(* Logix 5000 project; controller FV vendor 1 type 14 code 217 rev 31.11; software revision 31.00; part 22 of 63 *)
(* tags used below, declared in another part *)
   CheckTimeMask : INT;
   Delphi_Does_Eng_Func : BOOL;
   FR_FV29_AV04 : PlantItem;   // FV29_AV04
   FR_FV29_AV05 : PlantItem;   // FV29_AV05
   FR_FV29_AV06 : PlantItem;   // FV29_AV06
   FR_FV29_AV07 : PlantItem;   // FV29_AV07
   FR_N255 : INT[265];   // CHECKWORDS
   FR_VB2_AV01 : PlantItem;   // VB2_AV01
   FR_VB2_AV02 : PlantItem;   // VB2_AV02
   FR_VB2_AV03 : PlantItem;   // VB2_AV03
   FR_VB2_AV04 : PlantItem;   // VB2_AV04
   FR_VB2_AV05 : PlantItem;   // VB2_AV05
   FR_VB4_AV01 : PlantItem;   // VB4_AV01
   FR_VB4_AV02 : PlantItem;   // VB4_AV02
   FR_VB4_AV03 : PlantItem;   // VB4_AV03
   FR_VB4_AV04 : PlantItem;   // VB4_AV04
   TempChecktime : DINT;
(* FR_Common, continued *)

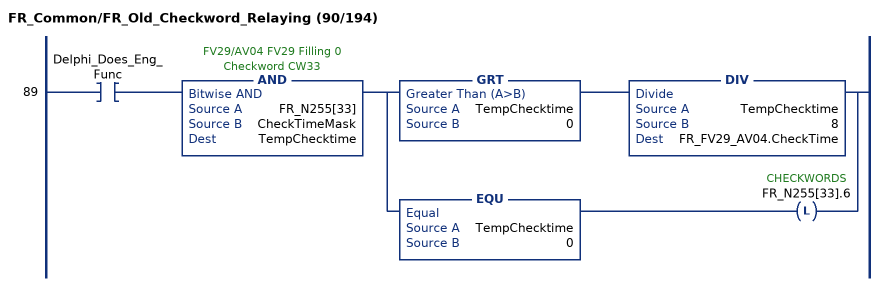
   [picture p394: FR_Common/FR_Old_Checkword_Relaying rungs 89-89]
   89: XIC(Delphi_Does_Eng_Func)AND(FR_N255[33],CheckTimeMask,TempChecktime)[GRT(TempChecktime,0) DIV(TempChecktime,8,FR_FV29_AV04.CheckTime) ,EQU(TempChecktime,0) OTL(FR_N255[33].6) ];
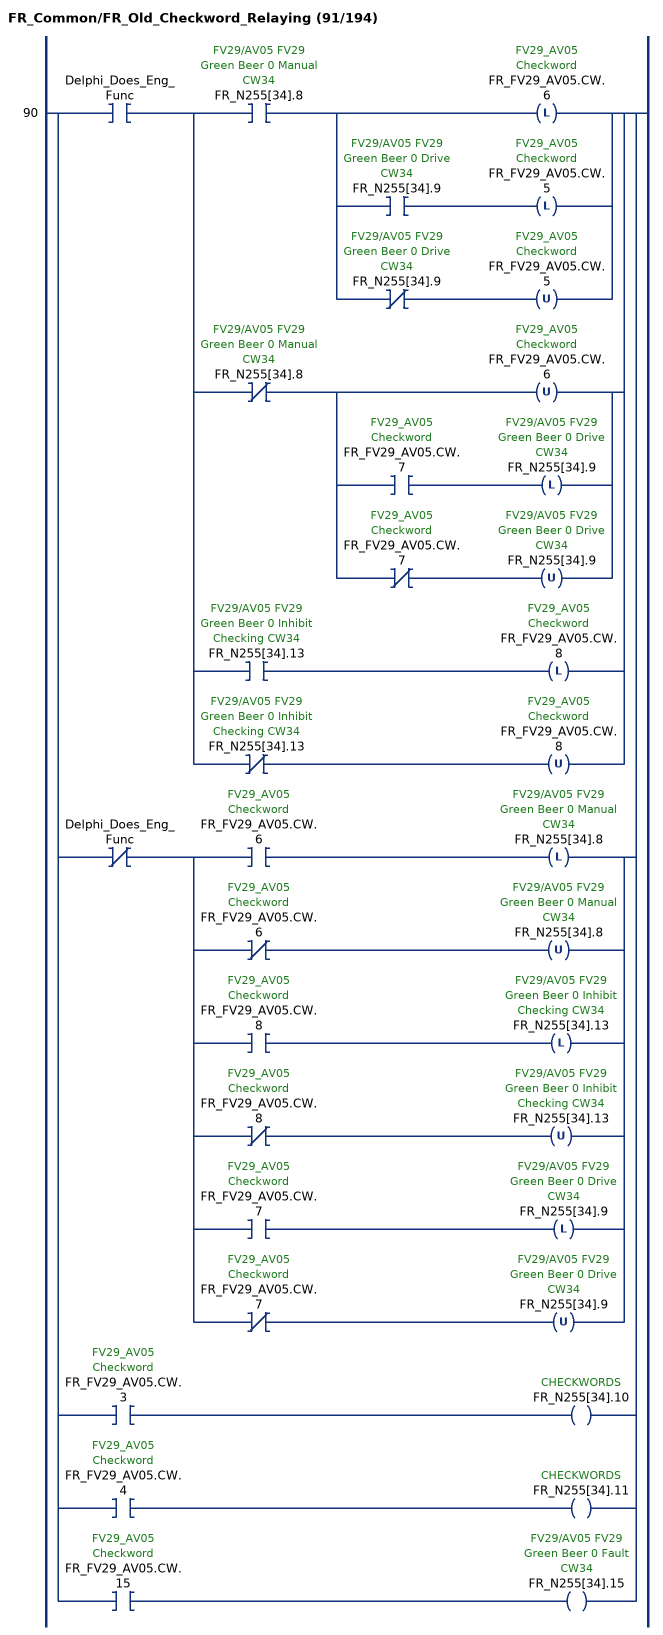
   90: [XIC(Delphi_Does_Eng_Func) [[XIC(FR_N255[34].8) [OTL(FR_FV29_AV05.CW.6) ,XIC(FR_N255[34].9) OTL(FR_FV29_AV05.CW.5) ,XIO(FR_N255[34].9) OTU(FR_FV29_AV05.CW.5) ] ,XIO(FR_N255[34].8) [OTU(FR_FV29_AV05.CW.6) ,[XIC(FR_FV29_AV05.CW.7) OTL(FR_N255[34].9) ,XIO(FR_FV29_AV05.CW.7) OTU(FR_N255[34].9) ] ] ] ,[XIC(FR_N255[34].13) OTL(FR_FV29_AV05.CW.8) ,XIO(FR_N255[34].13) OTU(FR_FV29_AV05.CW.8) ] ] ,XIO(Delphi_Does_Eng_Func) [[XIC(FR_FV29_AV05.CW.6) OTL(FR_N255[34].8) ,XIO(FR_FV29_AV05.CW.6) OTU(FR_N255[34].8) ] ,[XIC(FR_FV29_AV05.CW.8) OTL(FR_N255[34].13) ,XIO(FR_FV29_AV05.CW.8) OTU(FR_N255[34].13) ] ,[XIC(FR_FV29_AV05.CW.7) OTL(FR_N255[34].9) ,XIO(FR_FV29_AV05.CW.7) OTU(FR_N255[34].9) ] ] ,XIC(FR_FV29_AV05.CW.3) OTE(FR_N255[34].10) ,XIC(FR_FV29_AV05.CW.4) OTE(FR_N255[34].11) ,XIC(FR_FV29_AV05.CW.15) OTE(FR_N255[34].15) ];
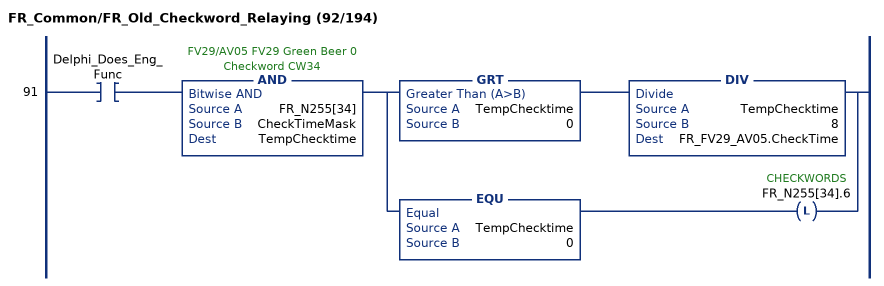
   91: XIC(Delphi_Does_Eng_Func)AND(FR_N255[34],CheckTimeMask,TempChecktime)[GRT(TempChecktime,0) DIV(TempChecktime,8,FR_FV29_AV05.CheckTime) ,EQU(TempChecktime,0) OTL(FR_N255[34].6) ];
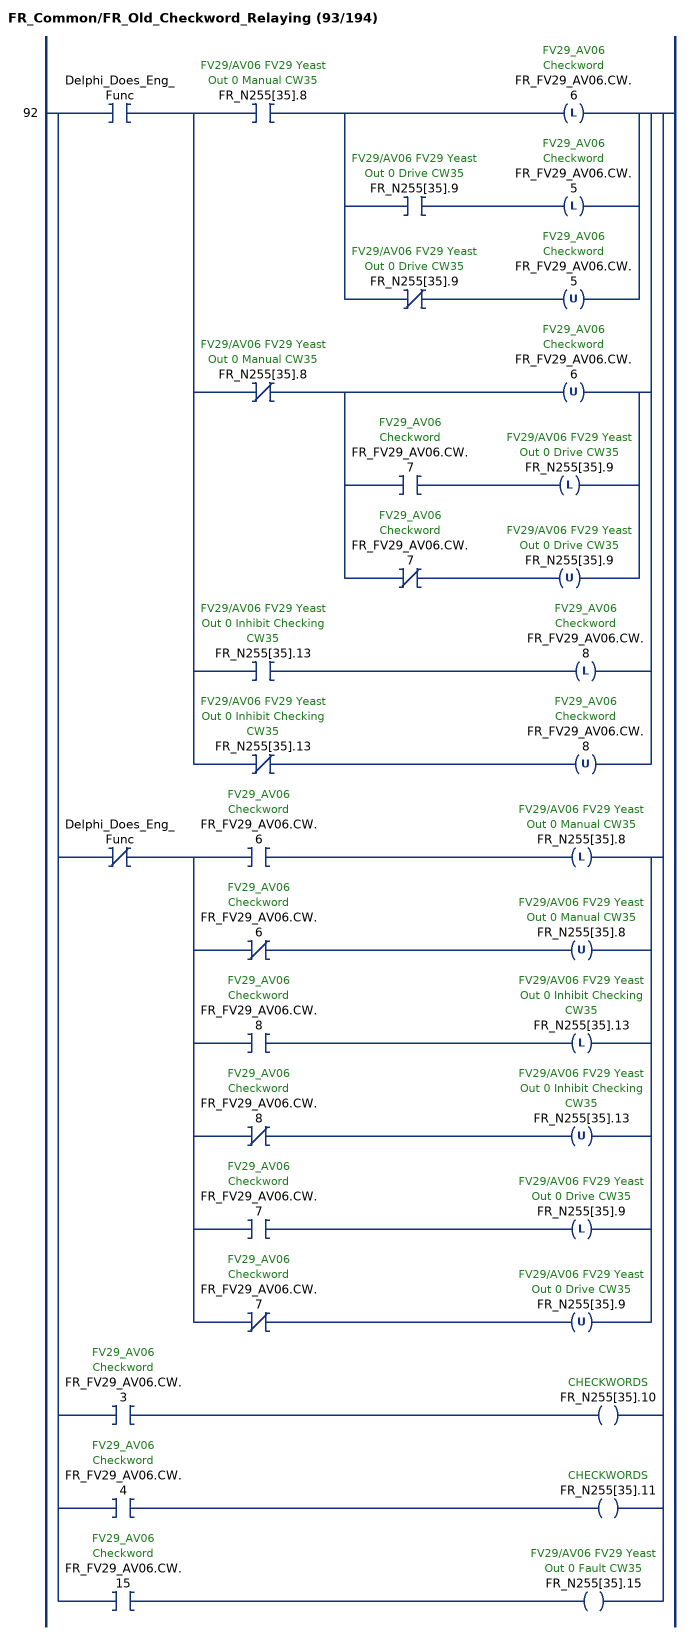
   92: [XIC(Delphi_Does_Eng_Func) [[XIC(FR_N255[35].8) [OTL(FR_FV29_AV06.CW.6) ,XIC(FR_N255[35].9) OTL(FR_FV29_AV06.CW.5) ,XIO(FR_N255[35].9) OTU(FR_FV29_AV06.CW.5) ] ,XIO(FR_N255[35].8) [OTU(FR_FV29_AV06.CW.6) ,[XIC(FR_FV29_AV06.CW.7) OTL(FR_N255[35].9) ,XIO(FR_FV29_AV06.CW.7) OTU(FR_N255[35].9) ] ] ] ,[XIC(FR_N255[35].13) OTL(FR_FV29_AV06.CW.8) ,XIO(FR_N255[35].13) OTU(FR_FV29_AV06.CW.8) ] ] ,XIO(Delphi_Does_Eng_Func) [[XIC(FR_FV29_AV06.CW.6) OTL(FR_N255[35].8) ,XIO(FR_FV29_AV06.CW.6) OTU(FR_N255[35].8) ] ,[XIC(FR_FV29_AV06.CW.8) OTL(FR_N255[35].13) ,XIO(FR_FV29_AV06.CW.8) OTU(FR_N255[35].13) ] ,[XIC(FR_FV29_AV06.CW.7) OTL(FR_N255[35].9) ,XIO(FR_FV29_AV06.CW.7) OTU(FR_N255[35].9) ] ] ,XIC(FR_FV29_AV06.CW.3) OTE(FR_N255[35].10) ,XIC(FR_FV29_AV06.CW.4) OTE(FR_N255[35].11) ,XIC(FR_FV29_AV06.CW.15) OTE(FR_N255[35].15) ];
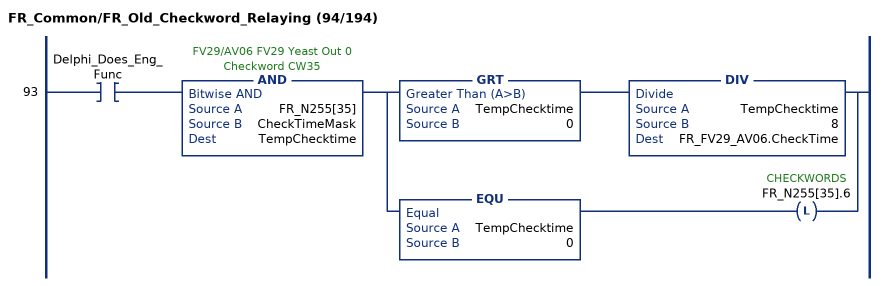
   93: XIC(Delphi_Does_Eng_Func)AND(FR_N255[35],CheckTimeMask,TempChecktime)[GRT(TempChecktime,0) DIV(TempChecktime,8,FR_FV29_AV06.CheckTime) ,EQU(TempChecktime,0) OTL(FR_N255[35].6) ];
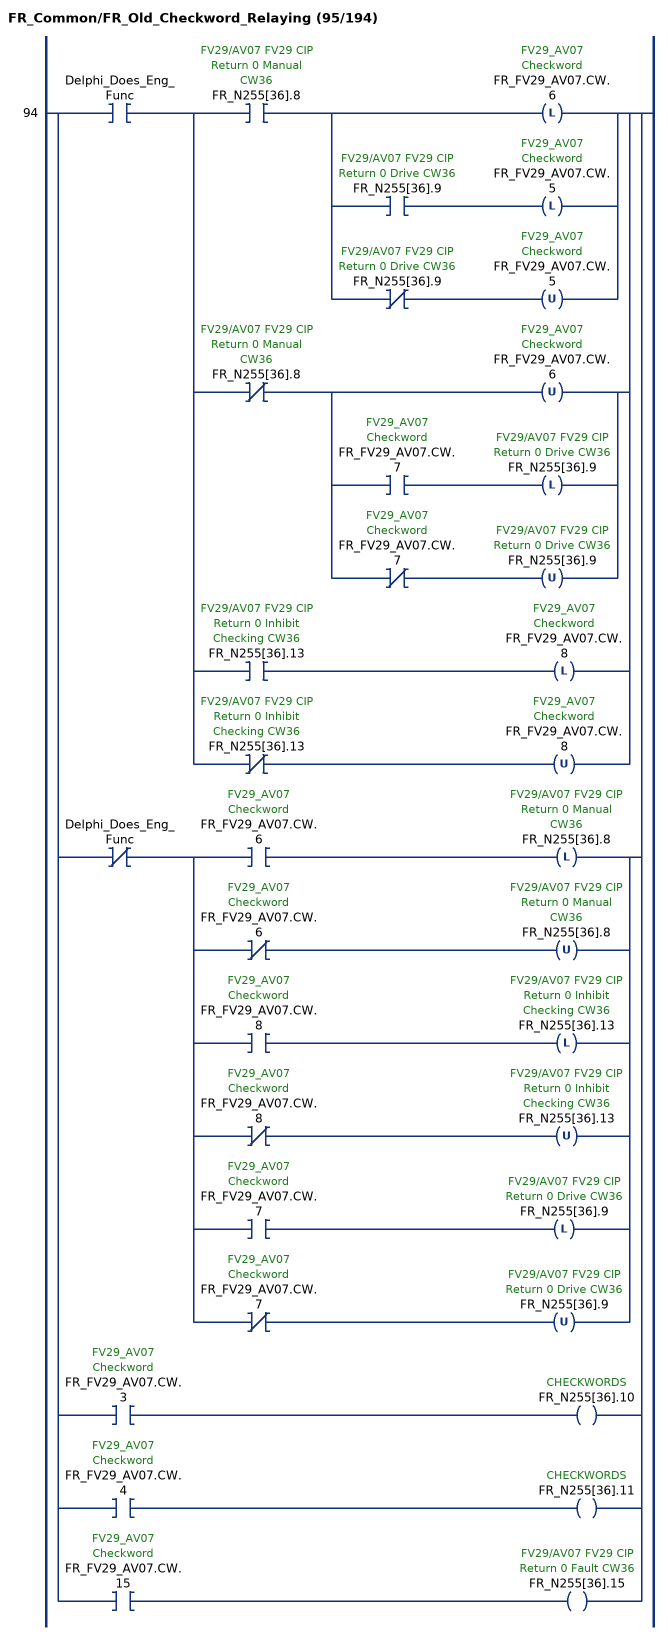
   94: [XIC(Delphi_Does_Eng_Func) [[XIC(FR_N255[36].8) [OTL(FR_FV29_AV07.CW.6) ,XIC(FR_N255[36].9) OTL(FR_FV29_AV07.CW.5) ,XIO(FR_N255[36].9) OTU(FR_FV29_AV07.CW.5) ] ,XIO(FR_N255[36].8) [OTU(FR_FV29_AV07.CW.6) ,[XIC(FR_FV29_AV07.CW.7) OTL(FR_N255[36].9) ,XIO(FR_FV29_AV07.CW.7) OTU(FR_N255[36].9) ] ] ] ,[XIC(FR_N255[36].13) OTL(FR_FV29_AV07.CW.8) ,XIO(FR_N255[36].13) OTU(FR_FV29_AV07.CW.8) ] ] ,XIO(Delphi_Does_Eng_Func) [[XIC(FR_FV29_AV07.CW.6) OTL(FR_N255[36].8) ,XIO(FR_FV29_AV07.CW.6) OTU(FR_N255[36].8) ] ,[XIC(FR_FV29_AV07.CW.8) OTL(FR_N255[36].13) ,XIO(FR_FV29_AV07.CW.8) OTU(FR_N255[36].13) ] ,[XIC(FR_FV29_AV07.CW.7) OTL(FR_N255[36].9) ,XIO(FR_FV29_AV07.CW.7) OTU(FR_N255[36].9) ] ] ,XIC(FR_FV29_AV07.CW.3) OTE(FR_N255[36].10) ,XIC(FR_FV29_AV07.CW.4) OTE(FR_N255[36].11) ,XIC(FR_FV29_AV07.CW.15) OTE(FR_N255[36].15) ];
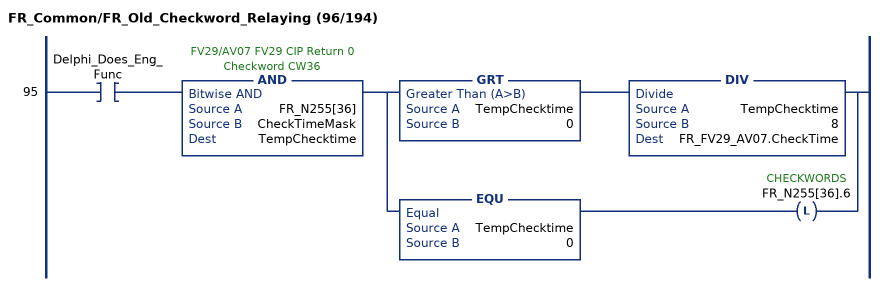
   95: XIC(Delphi_Does_Eng_Func)AND(FR_N255[36],CheckTimeMask,TempChecktime)[GRT(TempChecktime,0) DIV(TempChecktime,8,FR_FV29_AV07.CheckTime) ,EQU(TempChecktime,0) OTL(FR_N255[36].6) ];
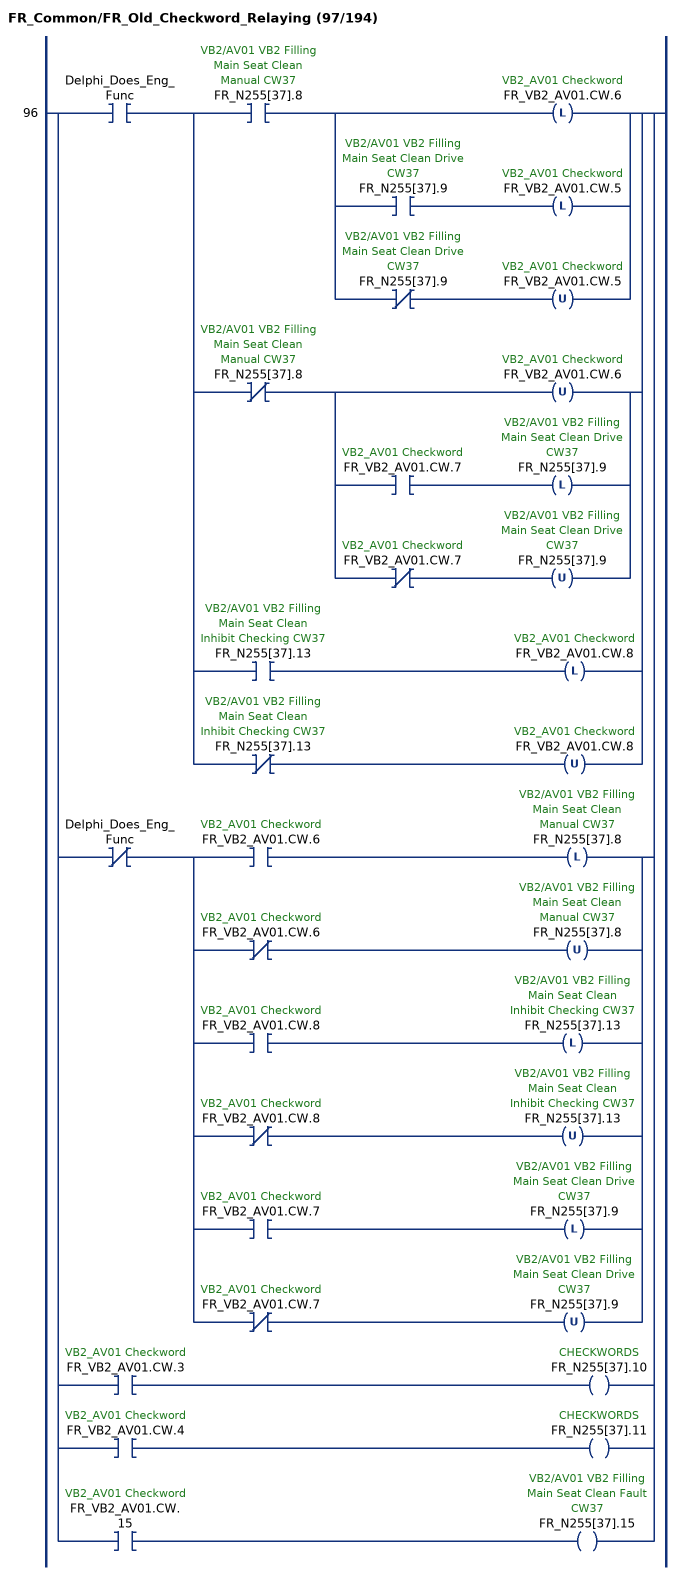
   96: [XIC(Delphi_Does_Eng_Func) [[XIC(FR_N255[37].8) [OTL(FR_VB2_AV01.CW.6) ,XIC(FR_N255[37].9) OTL(FR_VB2_AV01.CW.5) ,XIO(FR_N255[37].9) OTU(FR_VB2_AV01.CW.5) ] ,XIO(FR_N255[37].8) [OTU(FR_VB2_AV01.CW.6) ,[XIC(FR_VB2_AV01.CW.7) OTL(FR_N255[37].9) ,XIO(FR_VB2_AV01.CW.7) OTU(FR_N255[37].9) ] ] ] ,[XIC(FR_N255[37].13) OTL(FR_VB2_AV01.CW.8) ,XIO(FR_N255[37].13) OTU(FR_VB2_AV01.CW.8) ] ] ,XIO(Delphi_Does_Eng_Func) [[XIC(FR_VB2_AV01.CW.6) OTL(FR_N255[37].8) ,XIO(FR_VB2_AV01.CW.6) OTU(FR_N255[37].8) ] ,[XIC(FR_VB2_AV01.CW.8) OTL(FR_N255[37].13) ,XIO(FR_VB2_AV01.CW.8) OTU(FR_N255[37].13) ] ,[XIC(FR_VB2_AV01.CW.7) OTL(FR_N255[37].9) ,XIO(FR_VB2_AV01.CW.7) OTU(FR_N255[37].9) ] ] ,XIC(FR_VB2_AV01.CW.3) OTE(FR_N255[37].10) ,XIC(FR_VB2_AV01.CW.4) OTE(FR_N255[37].11) ,XIC(FR_VB2_AV01.CW.15) OTE(FR_N255[37].15) ];
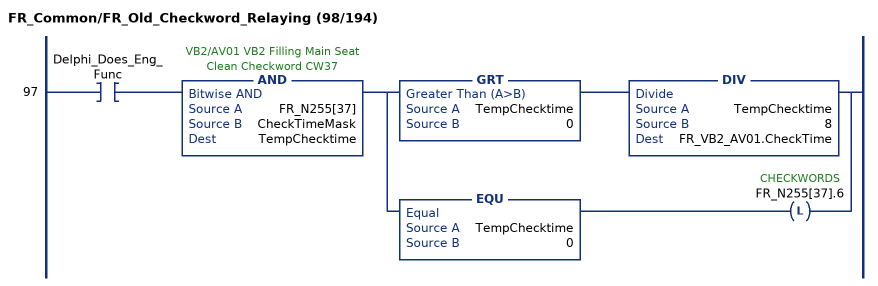
   97: XIC(Delphi_Does_Eng_Func)AND(FR_N255[37],CheckTimeMask,TempChecktime)[GRT(TempChecktime,0) DIV(TempChecktime,8,FR_VB2_AV01.CheckTime) ,EQU(TempChecktime,0) OTL(FR_N255[37].6) ];
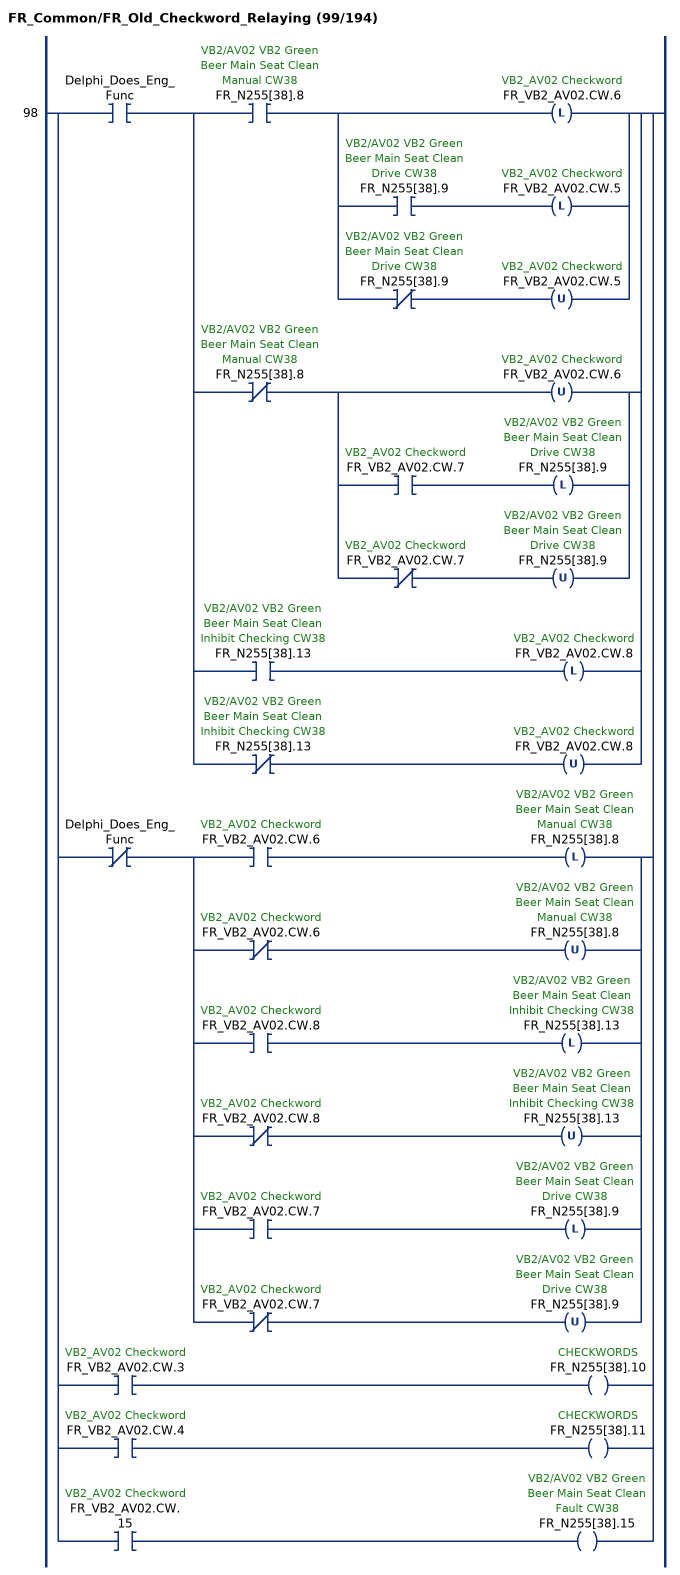
   98: [XIC(Delphi_Does_Eng_Func) [[XIC(FR_N255[38].8) [OTL(FR_VB2_AV02.CW.6) ,XIC(FR_N255[38].9) OTL(FR_VB2_AV02.CW.5) ,XIO(FR_N255[38].9) OTU(FR_VB2_AV02.CW.5) ] ,XIO(FR_N255[38].8) [OTU(FR_VB2_AV02.CW.6) ,[XIC(FR_VB2_AV02.CW.7) OTL(FR_N255[38].9) ,XIO(FR_VB2_AV02.CW.7) OTU(FR_N255[38].9) ] ] ] ,[XIC(FR_N255[38].13) OTL(FR_VB2_AV02.CW.8) ,XIO(FR_N255[38].13) OTU(FR_VB2_AV02.CW.8) ] ] ,XIO(Delphi_Does_Eng_Func) [[XIC(FR_VB2_AV02.CW.6) OTL(FR_N255[38].8) ,XIO(FR_VB2_AV02.CW.6) OTU(FR_N255[38].8) ] ,[XIC(FR_VB2_AV02.CW.8) OTL(FR_N255[38].13) ,XIO(FR_VB2_AV02.CW.8) OTU(FR_N255[38].13) ] ,[XIC(FR_VB2_AV02.CW.7) OTL(FR_N255[38].9) ,XIO(FR_VB2_AV02.CW.7) OTU(FR_N255[38].9) ] ] ,XIC(FR_VB2_AV02.CW.3) OTE(FR_N255[38].10) ,XIC(FR_VB2_AV02.CW.4) OTE(FR_N255[38].11) ,XIC(FR_VB2_AV02.CW.15) OTE(FR_N255[38].15) ];
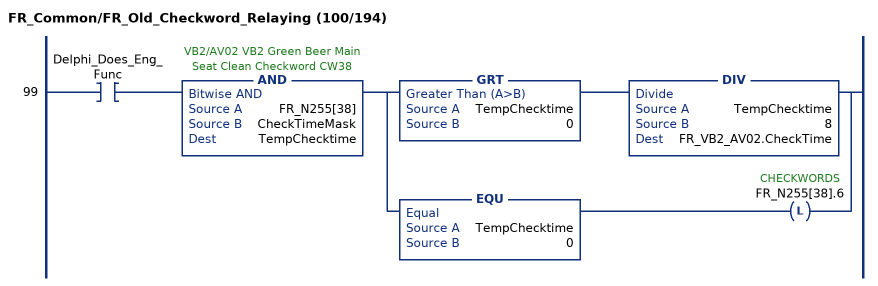
   99: XIC(Delphi_Does_Eng_Func)AND(FR_N255[38],CheckTimeMask,TempChecktime)[GRT(TempChecktime,0) DIV(TempChecktime,8,FR_VB2_AV02.CheckTime) ,EQU(TempChecktime,0) OTL(FR_N255[38].6) ];
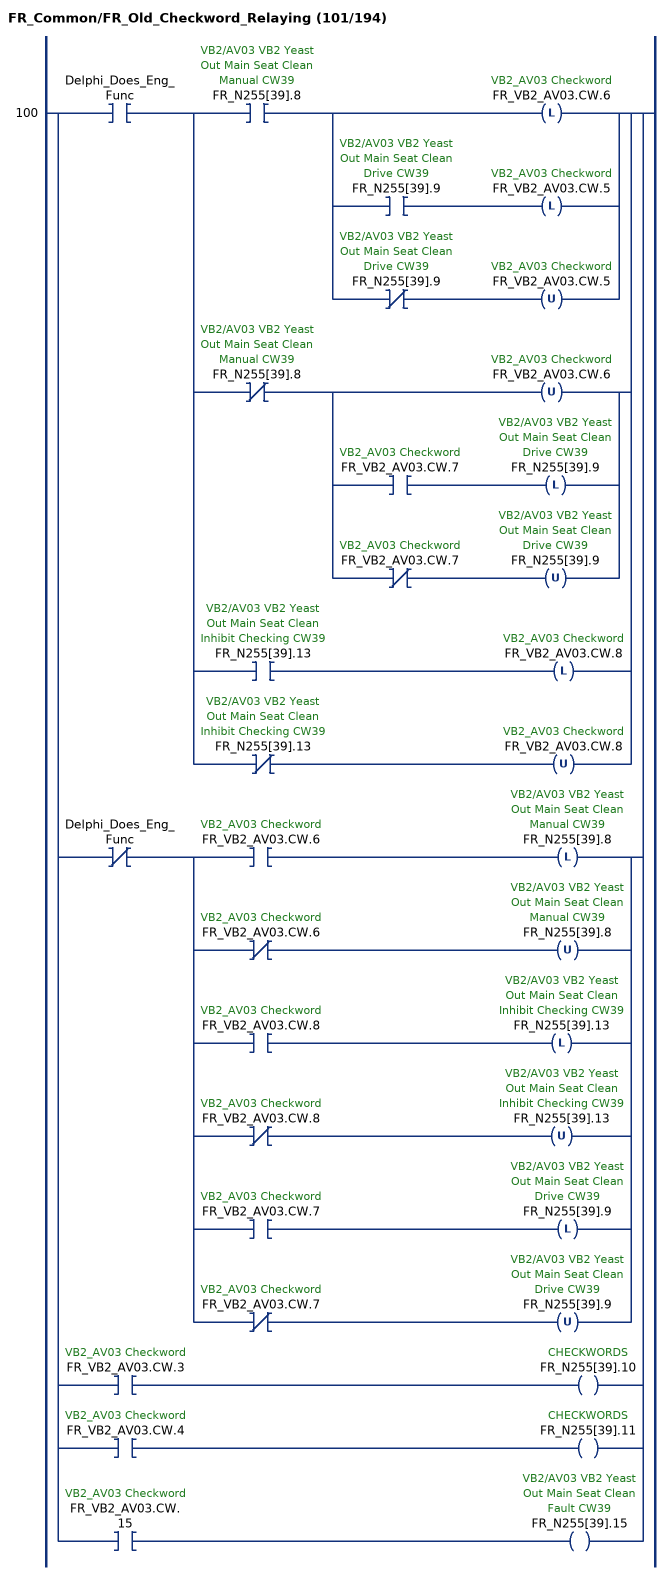
   100: [XIC(Delphi_Does_Eng_Func) [[XIC(FR_N255[39].8) [OTL(FR_VB2_AV03.CW.6) ,XIC(FR_N255[39].9) OTL(FR_VB2_AV03.CW.5) ,XIO(FR_N255[39].9) OTU(FR_VB2_AV03.CW.5) ] ,XIO(FR_N255[39].8) [OTU(FR_VB2_AV03.CW.6) ,[XIC(FR_VB2_AV03.CW.7) OTL(FR_N255[39].9) ,XIO(FR_VB2_AV03.CW.7) OTU(FR_N255[39].9) ] ] ] ,[XIC(FR_N255[39].13) OTL(FR_VB2_AV03.CW.8) ,XIO(FR_N255[39].13) OTU(FR_VB2_AV03.CW.8) ] ] ,XIO(Delphi_Does_Eng_Func) [[XIC(FR_VB2_AV03.CW.6) OTL(FR_N255[39].8) ,XIO(FR_VB2_AV03.CW.6) OTU(FR_N255[39].8) ] ,[XIC(FR_VB2_AV03.CW.8) OTL(FR_N255[39].13) ,XIO(FR_VB2_AV03.CW.8) OTU(FR_N255[39].13) ] ,[XIC(FR_VB2_AV03.CW.7) OTL(FR_N255[39].9) ,XIO(FR_VB2_AV03.CW.7) OTU(FR_N255[39].9) ] ] ,XIC(FR_VB2_AV03.CW.3) OTE(FR_N255[39].10) ,XIC(FR_VB2_AV03.CW.4) OTE(FR_N255[39].11) ,XIC(FR_VB2_AV03.CW.15) OTE(FR_N255[39].15) ];
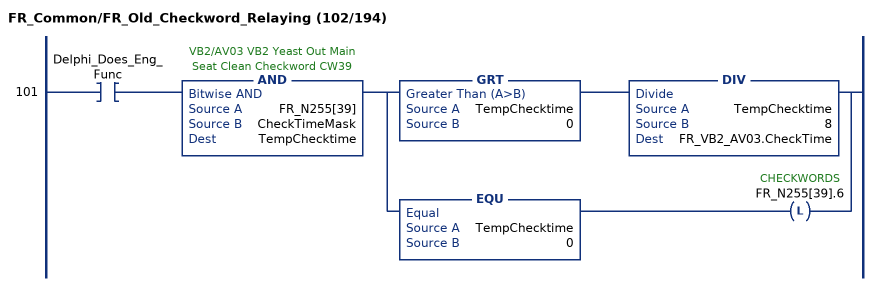
   101: XIC(Delphi_Does_Eng_Func)AND(FR_N255[39],CheckTimeMask,TempChecktime)[GRT(TempChecktime,0) DIV(TempChecktime,8,FR_VB2_AV03.CheckTime) ,EQU(TempChecktime,0) OTL(FR_N255[39].6) ];
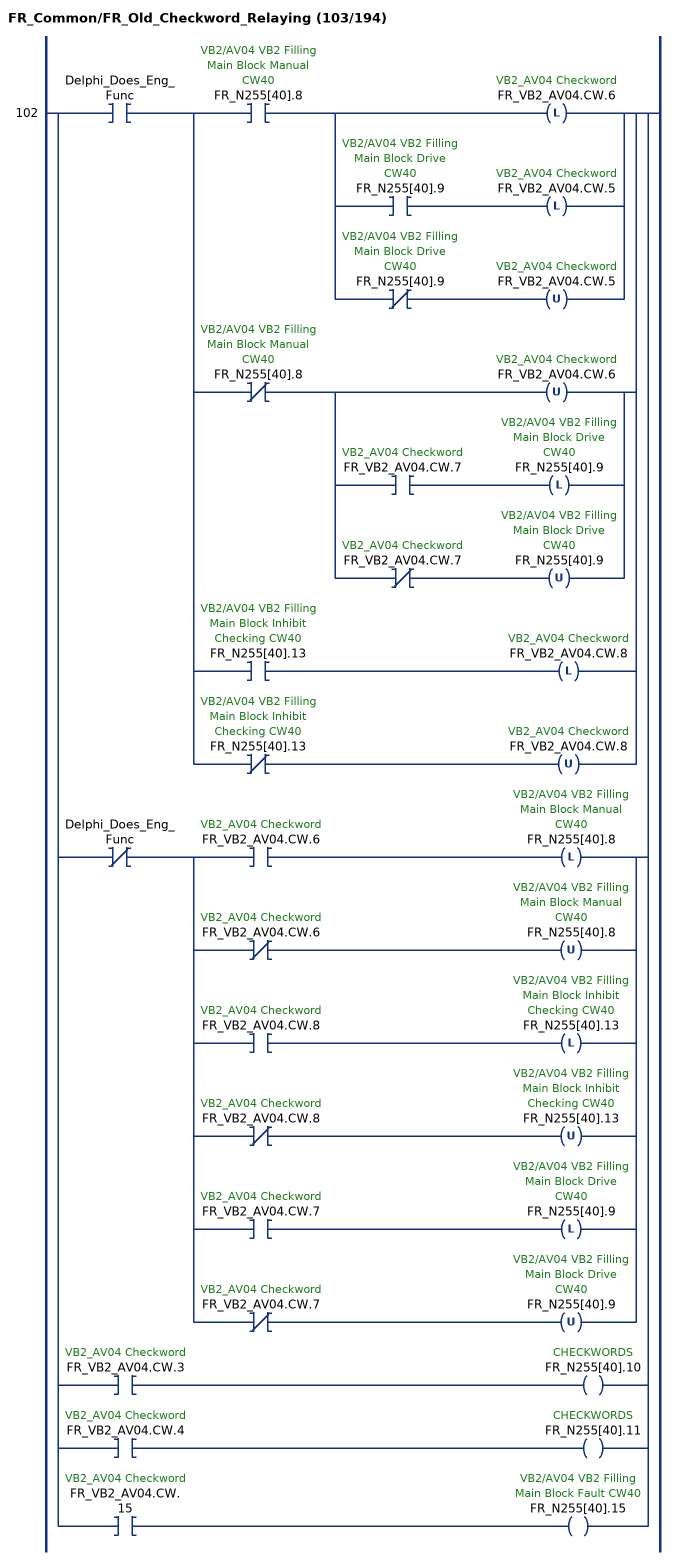
   102: [XIC(Delphi_Does_Eng_Func) [[XIC(FR_N255[40].8) [OTL(FR_VB2_AV04.CW.6) ,XIC(FR_N255[40].9) OTL(FR_VB2_AV04.CW.5) ,XIO(FR_N255[40].9) OTU(FR_VB2_AV04.CW.5) ] ,XIO(FR_N255[40].8) [OTU(FR_VB2_AV04.CW.6) ,[XIC(FR_VB2_AV04.CW.7) OTL(FR_N255[40].9) ,XIO(FR_VB2_AV04.CW.7) OTU(FR_N255[40].9) ] ] ] ,[XIC(FR_N255[40].13) OTL(FR_VB2_AV04.CW.8) ,XIO(FR_N255[40].13) OTU(FR_VB2_AV04.CW.8) ] ] ,XIO(Delphi_Does_Eng_Func) [[XIC(FR_VB2_AV04.CW.6) OTL(FR_N255[40].8) ,XIO(FR_VB2_AV04.CW.6) OTU(FR_N255[40].8) ] ,[XIC(FR_VB2_AV04.CW.8) OTL(FR_N255[40].13) ,XIO(FR_VB2_AV04.CW.8) OTU(FR_N255[40].13) ] ,[XIC(FR_VB2_AV04.CW.7) OTL(FR_N255[40].9) ,XIO(FR_VB2_AV04.CW.7) OTU(FR_N255[40].9) ] ] ,XIC(FR_VB2_AV04.CW.3) OTE(FR_N255[40].10) ,XIC(FR_VB2_AV04.CW.4) OTE(FR_N255[40].11) ,XIC(FR_VB2_AV04.CW.15) OTE(FR_N255[40].15) ];
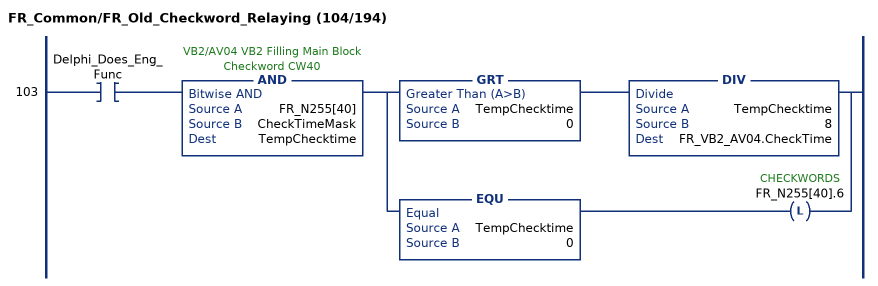
   103: XIC(Delphi_Does_Eng_Func)AND(FR_N255[40],CheckTimeMask,TempChecktime)[GRT(TempChecktime,0) DIV(TempChecktime,8,FR_VB2_AV04.CheckTime) ,EQU(TempChecktime,0) OTL(FR_N255[40].6) ];
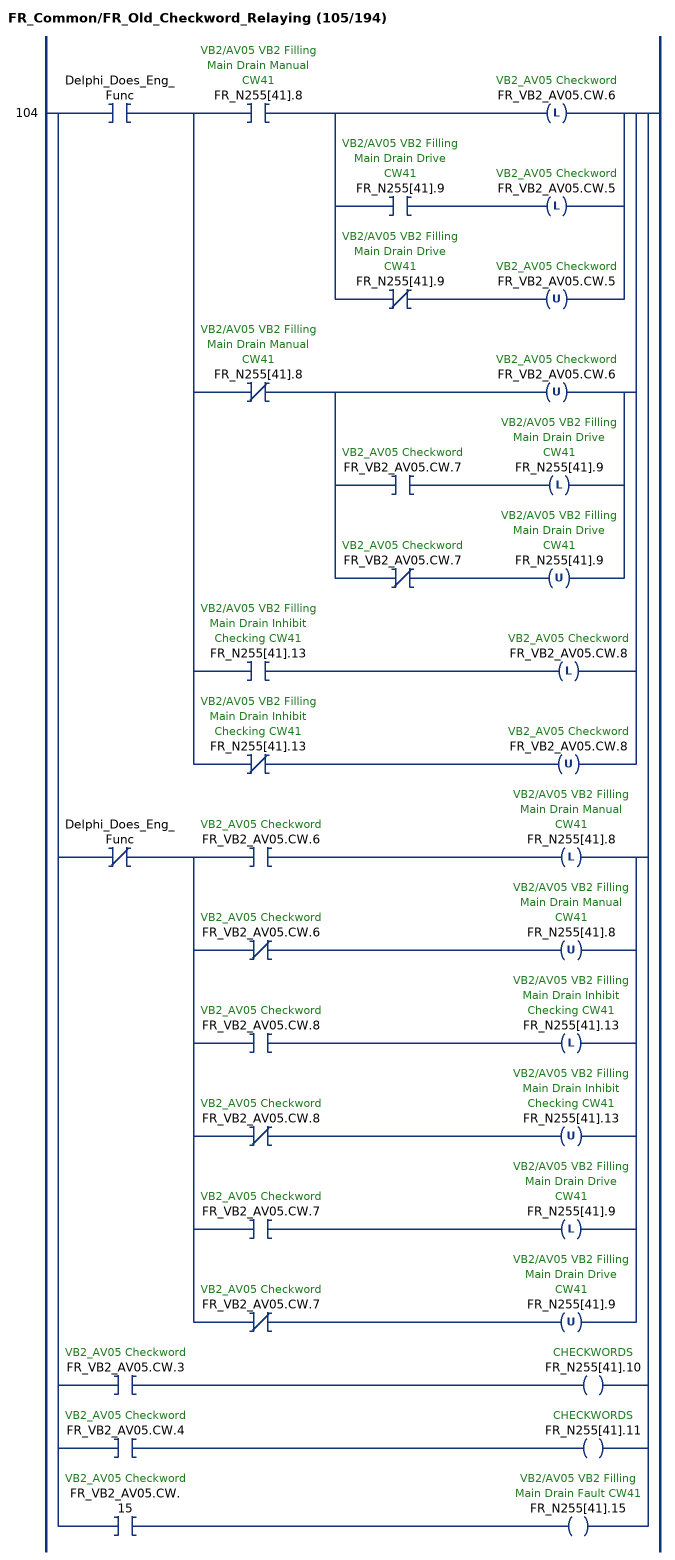
   104: [XIC(Delphi_Does_Eng_Func) [[XIC(FR_N255[41].8) [OTL(FR_VB2_AV05.CW.6) ,XIC(FR_N255[41].9) OTL(FR_VB2_AV05.CW.5) ,XIO(FR_N255[41].9) OTU(FR_VB2_AV05.CW.5) ] ,XIO(FR_N255[41].8) [OTU(FR_VB2_AV05.CW.6) ,[XIC(FR_VB2_AV05.CW.7) OTL(FR_N255[41].9) ,XIO(FR_VB2_AV05.CW.7) OTU(FR_N255[41].9) ] ] ] ,[XIC(FR_N255[41].13) OTL(FR_VB2_AV05.CW.8) ,XIO(FR_N255[41].13) OTU(FR_VB2_AV05.CW.8) ] ] ,XIO(Delphi_Does_Eng_Func) [[XIC(FR_VB2_AV05.CW.6) OTL(FR_N255[41].8) ,XIO(FR_VB2_AV05.CW.6) OTU(FR_N255[41].8) ] ,[XIC(FR_VB2_AV05.CW.8) OTL(FR_N255[41].13) ,XIO(FR_VB2_AV05.CW.8) OTU(FR_N255[41].13) ] ,[XIC(FR_VB2_AV05.CW.7) OTL(FR_N255[41].9) ,XIO(FR_VB2_AV05.CW.7) OTU(FR_N255[41].9) ] ] ,XIC(FR_VB2_AV05.CW.3) OTE(FR_N255[41].10) ,XIC(FR_VB2_AV05.CW.4) OTE(FR_N255[41].11) ,XIC(FR_VB2_AV05.CW.15) OTE(FR_N255[41].15) ];
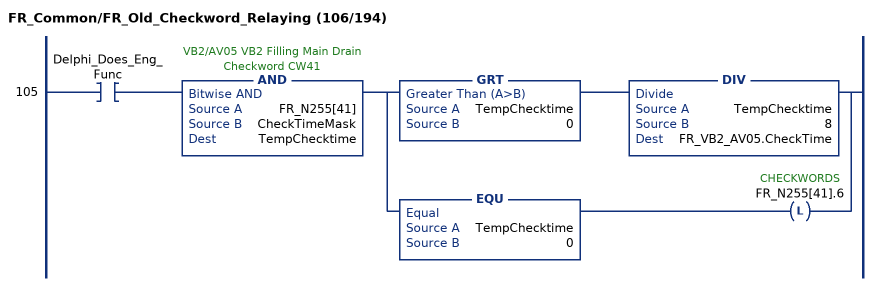
   105: XIC(Delphi_Does_Eng_Func)AND(FR_N255[41],CheckTimeMask,TempChecktime)[GRT(TempChecktime,0) DIV(TempChecktime,8,FR_VB2_AV05.CheckTime) ,EQU(TempChecktime,0) OTL(FR_N255[41].6) ];
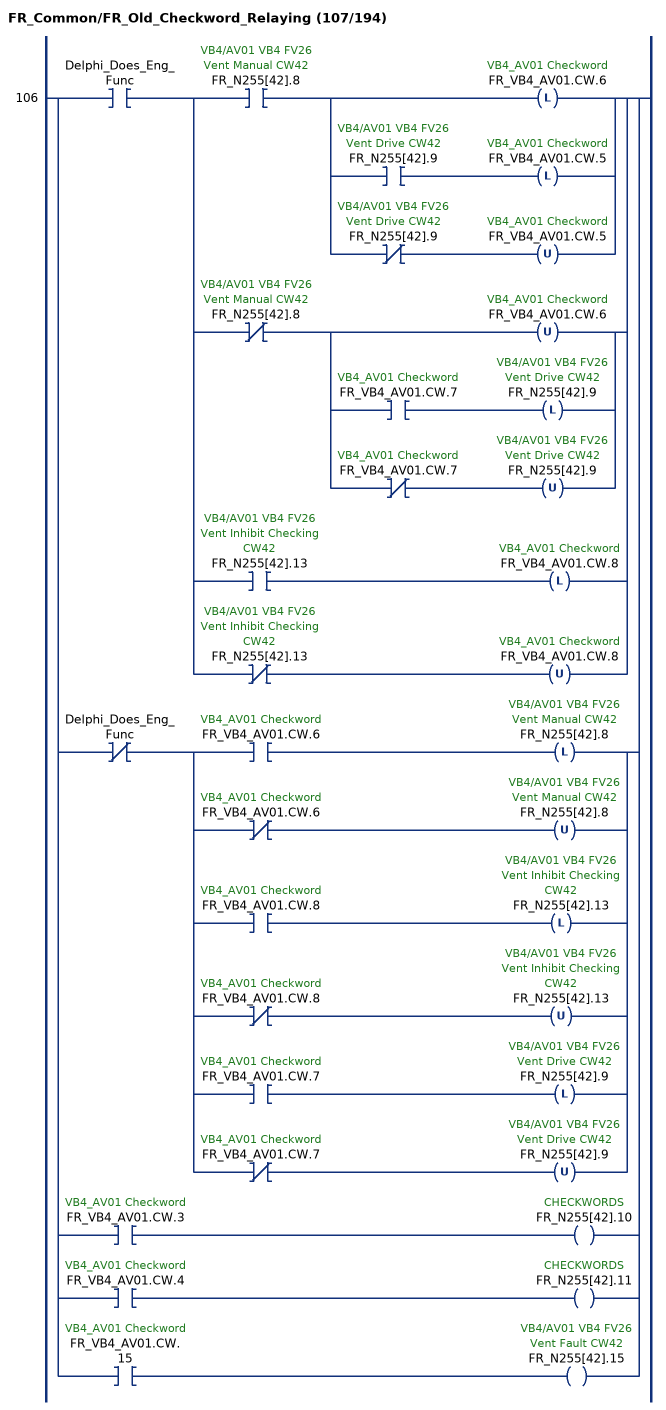
   106: [XIC(Delphi_Does_Eng_Func) [[XIC(FR_N255[42].8) [OTL(FR_VB4_AV01.CW.6) ,XIC(FR_N255[42].9) OTL(FR_VB4_AV01.CW.5) ,XIO(FR_N255[42].9) OTU(FR_VB4_AV01.CW.5) ] ,XIO(FR_N255[42].8) [OTU(FR_VB4_AV01.CW.6) ,[XIC(FR_VB4_AV01.CW.7) OTL(FR_N255[42].9) ,XIO(FR_VB4_AV01.CW.7) OTU(FR_N255[42].9) ] ] ] ,[XIC(FR_N255[42].13) OTL(FR_VB4_AV01.CW.8) ,XIO(FR_N255[42].13) OTU(FR_VB4_AV01.CW.8) ] ] ,XIO(Delphi_Does_Eng_Func) [[XIC(FR_VB4_AV01.CW.6) OTL(FR_N255[42].8) ,XIO(FR_VB4_AV01.CW.6) OTU(FR_N255[42].8) ] ,[XIC(FR_VB4_AV01.CW.8) OTL(FR_N255[42].13) ,XIO(FR_VB4_AV01.CW.8) OTU(FR_N255[42].13) ] ,[XIC(FR_VB4_AV01.CW.7) OTL(FR_N255[42].9) ,XIO(FR_VB4_AV01.CW.7) OTU(FR_N255[42].9) ] ] ,XIC(FR_VB4_AV01.CW.3) OTE(FR_N255[42].10) ,XIC(FR_VB4_AV01.CW.4) OTE(FR_N255[42].11) ,XIC(FR_VB4_AV01.CW.15) OTE(FR_N255[42].15) ];
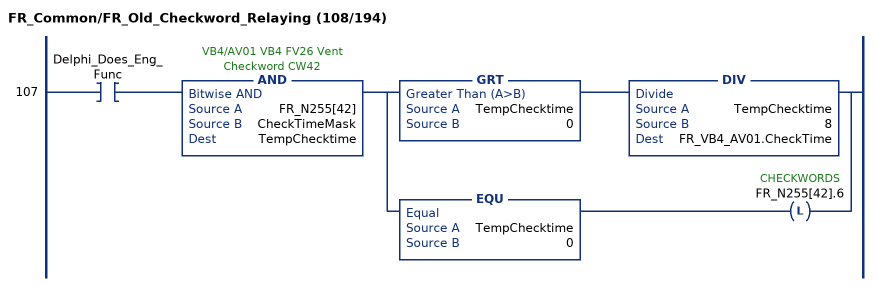
   107: XIC(Delphi_Does_Eng_Func)AND(FR_N255[42],CheckTimeMask,TempChecktime)[GRT(TempChecktime,0) DIV(TempChecktime,8,FR_VB4_AV01.CheckTime) ,EQU(TempChecktime,0) OTL(FR_N255[42].6) ];
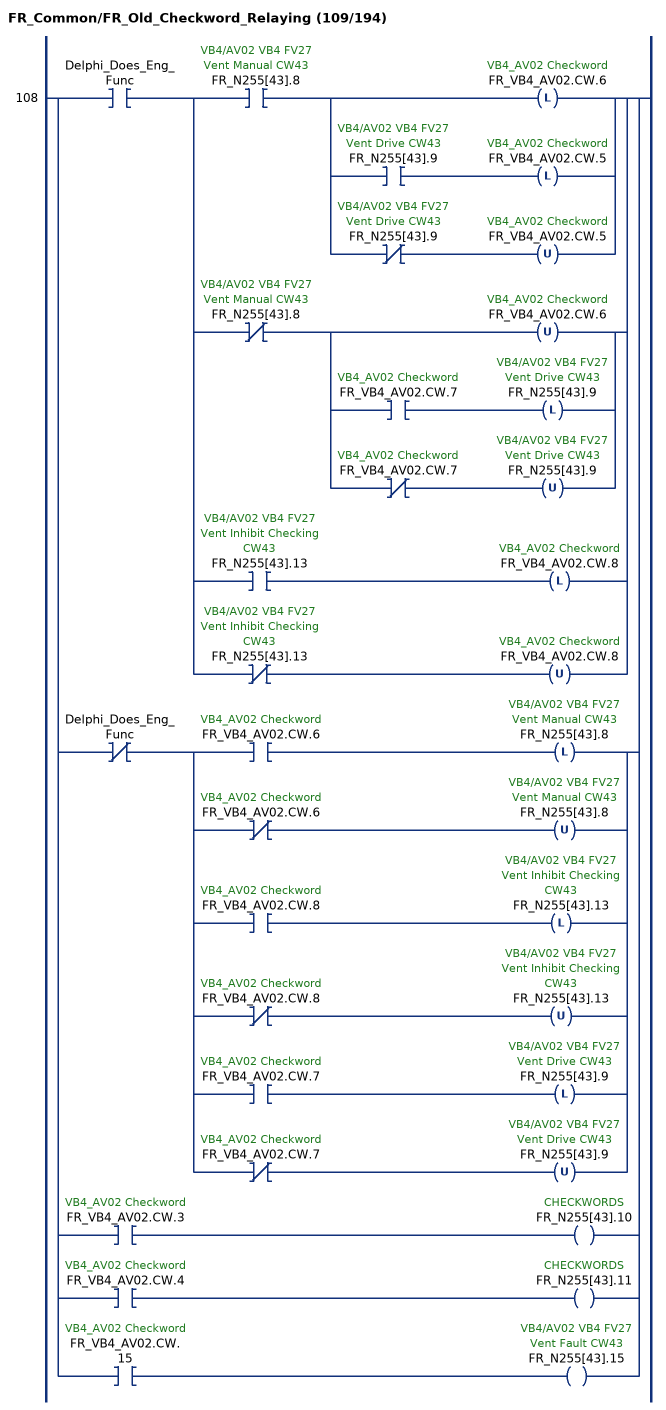
   108: [XIC(Delphi_Does_Eng_Func) [[XIC(FR_N255[43].8) [OTL(FR_VB4_AV02.CW.6) ,XIC(FR_N255[43].9) OTL(FR_VB4_AV02.CW.5) ,XIO(FR_N255[43].9) OTU(FR_VB4_AV02.CW.5) ] ,XIO(FR_N255[43].8) [OTU(FR_VB4_AV02.CW.6) ,[XIC(FR_VB4_AV02.CW.7) OTL(FR_N255[43].9) ,XIO(FR_VB4_AV02.CW.7) OTU(FR_N255[43].9) ] ] ] ,[XIC(FR_N255[43].13) OTL(FR_VB4_AV02.CW.8) ,XIO(FR_N255[43].13) OTU(FR_VB4_AV02.CW.8) ] ] ,XIO(Delphi_Does_Eng_Func) [[XIC(FR_VB4_AV02.CW.6) OTL(FR_N255[43].8) ,XIO(FR_VB4_AV02.CW.6) OTU(FR_N255[43].8) ] ,[XIC(FR_VB4_AV02.CW.8) OTL(FR_N255[43].13) ,XIO(FR_VB4_AV02.CW.8) OTU(FR_N255[43].13) ] ,[XIC(FR_VB4_AV02.CW.7) OTL(FR_N255[43].9) ,XIO(FR_VB4_AV02.CW.7) OTU(FR_N255[43].9) ] ] ,XIC(FR_VB4_AV02.CW.3) OTE(FR_N255[43].10) ,XIC(FR_VB4_AV02.CW.4) OTE(FR_N255[43].11) ,XIC(FR_VB4_AV02.CW.15) OTE(FR_N255[43].15) ];
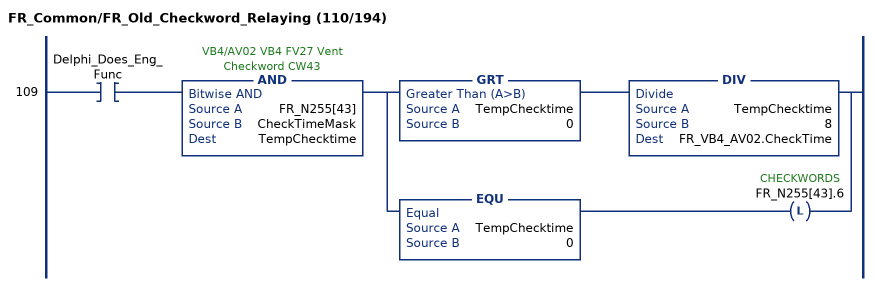
   109: XIC(Delphi_Does_Eng_Func)AND(FR_N255[43],CheckTimeMask,TempChecktime)[GRT(TempChecktime,0) DIV(TempChecktime,8,FR_VB4_AV02.CheckTime) ,EQU(TempChecktime,0) OTL(FR_N255[43].6) ];
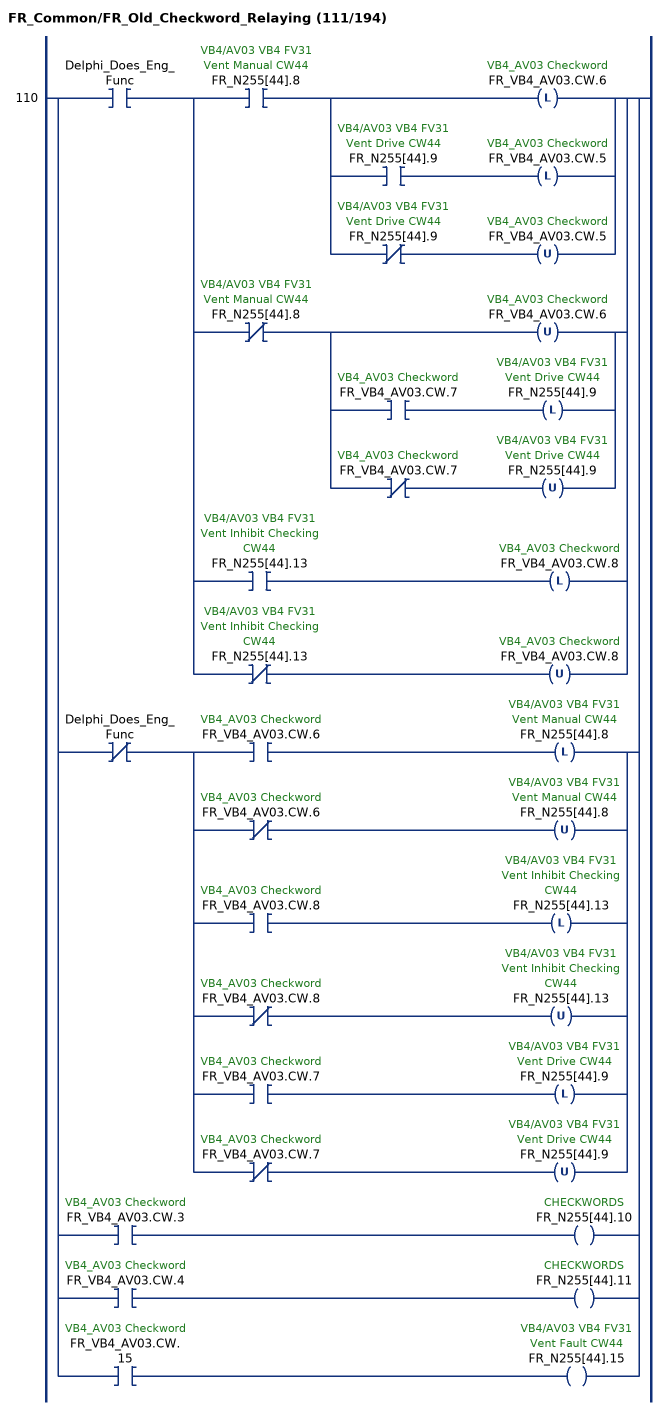
   110: [XIC(Delphi_Does_Eng_Func) [[XIC(FR_N255[44].8) [OTL(FR_VB4_AV03.CW.6) ,XIC(FR_N255[44].9) OTL(FR_VB4_AV03.CW.5) ,XIO(FR_N255[44].9) OTU(FR_VB4_AV03.CW.5) ] ,XIO(FR_N255[44].8) [OTU(FR_VB4_AV03.CW.6) ,[XIC(FR_VB4_AV03.CW.7) OTL(FR_N255[44].9) ,XIO(FR_VB4_AV03.CW.7) OTU(FR_N255[44].9) ] ] ] ,[XIC(FR_N255[44].13) OTL(FR_VB4_AV03.CW.8) ,XIO(FR_N255[44].13) OTU(FR_VB4_AV03.CW.8) ] ] ,XIO(Delphi_Does_Eng_Func) [[XIC(FR_VB4_AV03.CW.6) OTL(FR_N255[44].8) ,XIO(FR_VB4_AV03.CW.6) OTU(FR_N255[44].8) ] ,[XIC(FR_VB4_AV03.CW.8) OTL(FR_N255[44].13) ,XIO(FR_VB4_AV03.CW.8) OTU(FR_N255[44].13) ] ,[XIC(FR_VB4_AV03.CW.7) OTL(FR_N255[44].9) ,XIO(FR_VB4_AV03.CW.7) OTU(FR_N255[44].9) ] ] ,XIC(FR_VB4_AV03.CW.3) OTE(FR_N255[44].10) ,XIC(FR_VB4_AV03.CW.4) OTE(FR_N255[44].11) ,XIC(FR_VB4_AV03.CW.15) OTE(FR_N255[44].15) ];
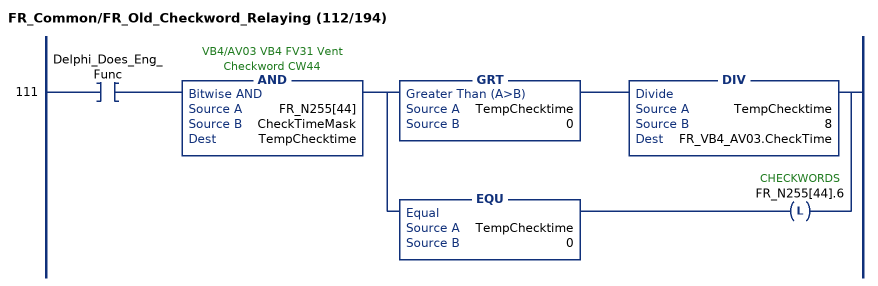
   111: XIC(Delphi_Does_Eng_Func)AND(FR_N255[44],CheckTimeMask,TempChecktime)[GRT(TempChecktime,0) DIV(TempChecktime,8,FR_VB4_AV03.CheckTime) ,EQU(TempChecktime,0) OTL(FR_N255[44].6) ];
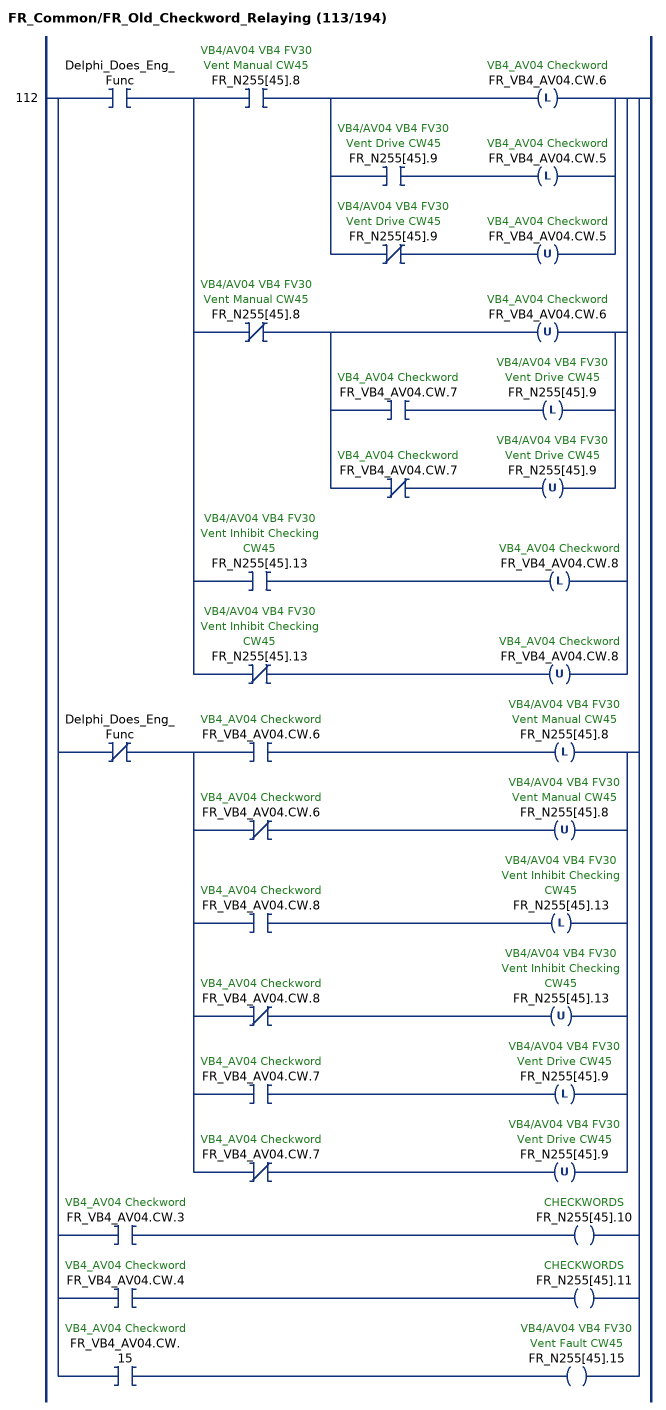
   112: [XIC(Delphi_Does_Eng_Func) [[XIC(FR_N255[45].8) [OTL(FR_VB4_AV04.CW.6) ,XIC(FR_N255[45].9) OTL(FR_VB4_AV04.CW.5) ,XIO(FR_N255[45].9) OTU(FR_VB4_AV04.CW.5) ] ,XIO(FR_N255[45].8) [OTU(FR_VB4_AV04.CW.6) ,[XIC(FR_VB4_AV04.CW.7) OTL(FR_N255[45].9) ,XIO(FR_VB4_AV04.CW.7) OTU(FR_N255[45].9) ] ] ] ,[XIC(FR_N255[45].13) OTL(FR_VB4_AV04.CW.8) ,XIO(FR_N255[45].13) OTU(FR_VB4_AV04.CW.8) ] ] ,XIO(Delphi_Does_Eng_Func) [[XIC(FR_VB4_AV04.CW.6) OTL(FR_N255[45].8) ,XIO(FR_VB4_AV04.CW.6) OTU(FR_N255[45].8) ] ,[XIC(FR_VB4_AV04.CW.8) OTL(FR_N255[45].13) ,XIO(FR_VB4_AV04.CW.8) OTU(FR_N255[45].13) ] ,[XIC(FR_VB4_AV04.CW.7) OTL(FR_N255[45].9) ,XIO(FR_VB4_AV04.CW.7) OTU(FR_N255[45].9) ] ] ,XIC(FR_VB4_AV04.CW.3) OTE(FR_N255[45].10) ,XIC(FR_VB4_AV04.CW.4) OTE(FR_N255[45].11) ,XIC(FR_VB4_AV04.CW.15) OTE(FR_N255[45].15) ];
